// TIA Portal project "Project2_Pompe" (V15.1)

(* hardware
DEVICE "S71500/ET200MP station_1"  S7-1500 station
   slot 0: "Rail_0"  Rack  6ES7 590-1***0-0AA0
   slot 1: "PLC_1"  CPU 1513-1 PN  6ES7 513-1AL02-0AB0  V2.6
      slot 3: "CPU display_1"  6ES7591-1AA00-0AA0
DEVICE "HMI_1"  KTP900 Basic PN
   slot 0: "HMI_1"  KTP900 Basic PN  6AV2 123-2JB03-0AX0  15.1.0.0
   slot 1: "HMI_RT_1"  KTP900 Basic PN  6AV2 123-2JB03-0AX0  15.1.0.0
   slot 5: "HMI_1.IE_CP_1"  PROFINET Interface  15.0.1.0
      slot 1: "PROFINET Interface_1"  PROFINET Interface
         slot 1: "Port_1"  Port
*)

// ===== PLC "PLC_1"  CPU 1513-1 PN =====

VAR_GLOBAL   // PLC tag table "Default tag table"
   "Clock_Byte" AT %MB0 : Byte;
   "Clock_10Hz" AT %M0.0 : Bool;
   "Clock_5Hz" AT %M0.1 : Bool;
   "Clock_2.5Hz" AT %M0.2 : Bool;
   "Clock_2Hz" AT %M0.3 : Bool;
   "Clock_1.25Hz" AT %M0.4 : Bool;
   "Clock_1Hz" AT %M0.5 : Bool;
   "Clock_0.625Hz" AT %M0.6 : Bool;
   "Clock_0.5Hz" AT %M0.7 : Bool;
END_VAR

VAR_GLOBAL   // PLC tag table "Intrari"
   "S1(clk)" AT %I0.0 : Bool;
   "S2(ctrclk)" AT %I0.1 : Bool;
   "s0(stop)" AT %I0.2 : Bool;
   "ptc(esd)" AT %I0.3 : Bool;
   "ss" AT %I0.4 : Bool;
END_VAR

VAR_GLOBAL   // PLC tag table "Iesiri"
   "K1(clk)" AT %Q0.0 : Bool;
   "K2(ctrclk)" AT %Q0.1 : Bool;
   "K3(triunghi)" AT %Q0.2 : Bool;
   "K4(stea)" AT %Q0.3 : Bool;
END_VAR

VAR_GLOBAL   // PLC tag table "Auxiliare"
   "M_pornit" AT %M1.0 : Bool;
   "passed_k3" AT %M1.1 : Bool;
   "reset urgenta" AT %M1.2 : Bool;
   "temporizare K4" AT %M1.3 : Bool;
   "permisie start" AT %M1.4 : Bool;
   "urgenta bit" AT %M1.5 : Bool;
END_VAR

// folder: System blocks/Program resources

DATA_BLOCK "IEC_Timer_0_DB"   // DB1
{ S7_Optimized_Access := 'TRUE' }
AUTHOR : Simatic
FAMILY : IEC
NAME : IEC_TMR
VERSION : 1.0
// stored: InstanceOfName IEC_TIMER
"IEC_TIMER"
BEGIN
END_DATA_BLOCK

DATA_BLOCK "IEC_Timer_0_DB_1"   // DB2
{ S7_Optimized_Access := 'TRUE' }
AUTHOR : Simatic
FAMILY : IEC
NAME : IEC_TMR
VERSION : 1.0
// stored: InstanceOfName IEC_TIMER
"IEC_TIMER"
BEGIN
END_DATA_BLOCK

// folder: (top level)

FUNCTION_BLOCK "Block_1"   // FB1, LAD
{ S7_Optimized_Access := 'TRUE' }
VERSION : 0.1
   VAR_INPUT
      start : Bool;
      stop : Bool;
      ESD : Bool;
   END_VAR
   VAR_OUTPUT
      "comanda motor" : Bool;
   END_VAR
BEGIN

REGION Network 1
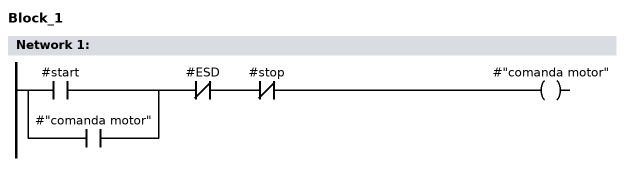
   RUNG wire#powerrail
      Contact( #start )
      wire#w1
      I_Contact( #ESD )
      I_Contact( #stop )
      Coil( #"comanda motor" )
   END_RUNG
   RUNG wire#powerrail
      Contact( #"comanda motor" )
   END_RUNG wire#w1
   // the same network as SCL:
   #"comanda motor" := (#start OR #"comanda motor") AND NOT #ESD AND NOT #stop;
END_REGION
END_FUNCTION_BLOCK

ORGANIZATION_BLOCK "Main"   // OB1, LAD, ProgramCycle
TITLE = "Main Program Sweep (Cycle)"
{ S7_Optimized_Access := 'TRUE' }
VERSION : 0.1
   VAR_INPUT
      Initial_Call : Bool;   // Initial call of this OB
      Remanence : Bool;   // =True, if remanent data are available
   END_VAR
BEGIN

REGION Network 1: selecteaza pe ce directie sa porneasca
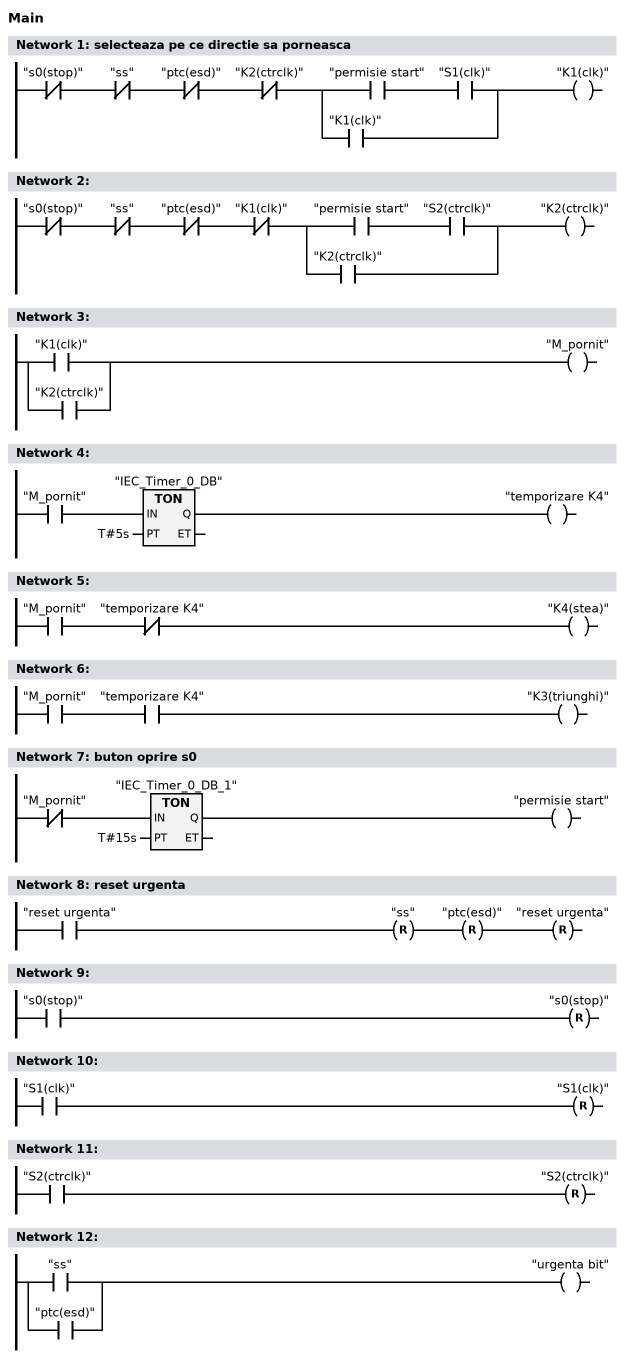
   RUNG wire#powerrail
      I_Contact( "s0(stop)" )
      I_Contact( "ss" )
      I_Contact( "ptc(esd)" )
      I_Contact( "K2(ctrclk)" )
      wire#w1
      Contact( "permisie start" )
      Contact( "S1(clk)" )
      wire#w2
      Coil( "K1(clk)" )
   END_RUNG
   RUNG wire#w1
      Contact( "K1(clk)" )
   END_RUNG wire#w2
   // the same network as SCL:
   "K1(clk)" := NOT "s0(stop)" AND NOT "ss" AND NOT "ptc(esd)" AND NOT "K2(ctrclk)" AND (("permisie start" AND "S1(clk)") OR "K1(clk)");
END_REGION

REGION Network 2
   RUNG wire#powerrail
      I_Contact( "s0(stop)" )
      I_Contact( "ss" )
      I_Contact( "ptc(esd)" )
      I_Contact( "K1(clk)" )
      wire#w1
      Contact( "permisie start" )
      Contact( "S2(ctrclk)" )
      wire#w2
      Coil( "K2(ctrclk)" )
   END_RUNG
   RUNG wire#w1
      Contact( "K2(ctrclk)" )
   END_RUNG wire#w2
   // the same network as SCL:
   "K2(ctrclk)" := NOT "s0(stop)" AND NOT "ss" AND NOT "ptc(esd)" AND NOT "K1(clk)" AND (("permisie start" AND "S2(ctrclk)") OR "K2(ctrclk)");
END_REGION

REGION Network 3
   RUNG wire#powerrail
      Contact( "K1(clk)" )
      wire#w1
      Coil( "M_pornit" )
   END_RUNG
   RUNG wire#powerrail
      Contact( "K2(ctrclk)" )
   END_RUNG wire#w1
   // the same network as SCL:
   "M_pornit" := "K1(clk)" OR "K2(ctrclk)";
END_REGION

REGION Network 4
   "IEC_Timer_0_DB".TON(IN := "M_pornit", PT := T#5s);
   "temporizare K4" := "IEC_Timer_0_DB".Q;
END_REGION

REGION Network 5
   RUNG wire#powerrail
      Contact( "M_pornit" )
      I_Contact( "temporizare K4" )
      Coil( "K4(stea)" )
   END_RUNG
   // the same network as SCL:
   "K4(stea)" := "M_pornit" AND NOT "temporizare K4";
END_REGION

REGION Network 6
   RUNG wire#powerrail
      Contact( "M_pornit" )
      Contact( "temporizare K4" )
      Coil( "K3(triunghi)" )
   END_RUNG
   // the same network as SCL:
   "K3(triunghi)" := "M_pornit" AND "temporizare K4";
END_REGION

REGION Network 7: buton oprire s0
   "IEC_Timer_0_DB_1".TON(IN := NOT "M_pornit", PT := T#15s);
   "permisie start" := "IEC_Timer_0_DB_1".Q;
END_REGION

REGION Network 8: reset urgenta
   RUNG wire#powerrail
      Contact( "reset urgenta" )
      R_Coil( "ss" )
      R_Coil( "ptc(esd)" )
      R_Coil( "reset urgenta" )
   END_RUNG
   // the same network as SCL:
   IF "reset urgenta" THEN
       "ss" := FALSE;
       "ptc(esd)" := FALSE;
       "reset urgenta" := FALSE;
   END_IF;
END_REGION

REGION Network 9
   RUNG wire#powerrail
      Contact( "s0(stop)" )
      R_Coil( "s0(stop)" )
   END_RUNG
   // the same network as SCL:
   IF "s0(stop)" THEN "s0(stop)" := FALSE; END_IF;
END_REGION

REGION Network 10
   RUNG wire#powerrail
      Contact( "S1(clk)" )
      R_Coil( "S1(clk)" )
   END_RUNG
   // the same network as SCL:
   IF "S1(clk)" THEN "S1(clk)" := FALSE; END_IF;
END_REGION

REGION Network 11
   RUNG wire#powerrail
      Contact( "S2(ctrclk)" )
      R_Coil( "S2(ctrclk)" )
   END_RUNG
   // the same network as SCL:
   IF "S2(ctrclk)" THEN "S2(ctrclk)" := FALSE; END_IF;
END_REGION

REGION Network 12
   RUNG wire#powerrail
      Contact( "ss" )
      wire#w1
      Coil( "urgenta bit" )
   END_RUNG
   RUNG wire#powerrail
      Contact( "ptc(esd)" )
   END_RUNG wire#w1
   // the same network as SCL:
   "urgenta bit" := "ss" OR "ptc(esd)";
END_REGION
END_ORGANIZATION_BLOCK

(* ===== HMI "HMI_RT_1" =====
system functions are stored by id; their names below are inferred from use
connection "HMI_Connection_1": ETHERNET, SMART_S7_1500_OMS

HMI tags "Default tag table"
   "Tag_ScreenNumber" : UInt, internal
   "s0(stop)" : Bool = PLC "s0(stop)" AT %I0.2, 1 s
   "S1(clk)" : Bool = PLC "S1(clk)" AT %I0.0, 1 s
   "S2(ctrclk)" : Bool = PLC "S2(ctrclk)" AT %I0.1, 1 s
   "IEC_Timer_0_DB_1_ET" : Time = PLC IEC_Timer_0_DB_1.ET, 1 s
   "IEC_Timer_0_DB_ET" : Time = PLC IEC_Timer_0_DB.ET, 1 s
   "K1(clk)" : Bool = PLC "K1(clk)" AT %Q0.0, 1 s
   "K2(ctrclk)" : Bool = PLC "K2(ctrclk)" AT %Q0.1, 1 s
   "K3(triunghi)" : Bool = PLC "K3(triunghi)" AT %Q0.2, 1 s
   "K4(stea)" : Bool = PLC "K4(stea)" AT %Q0.3, 1 s
   "ss" : Bool = PLC ss AT %I0.4, 1 s
   "M_pornit" : Bool = PLC M_pornit AT %M1.0, 1 s
   "reset urgenta" : Bool = PLC "reset urgenta" AT %M1.2, 1 s
   "ptc(esd)" : Bool = PLC "ptc(esd)" AT %I0.3, 1 s
   "urgenta bit" : Bool = PLC "urgenta bit" AT %M1.5, 1 s

Template "Template_1" 800x480
   Button "Exit" at 722,440 size 55x39; TextOff 'Exit'; PictureOff "ExitRuntime_KTP900_Basic_PN_TR"; PictureOn "ExitRuntime_KTP900_Basic_PN_TR"
      on Release: StopRuntime(0)
   Button "Template_Button" at 622,440 size 55x39; TextOff 'Text'
   Button "Template_Button_1" at 522,440 size 55x39; TextOff 'Text'
   Button "Template_Button_2" at 422,440 size 55x39; TextOff 'Text'
   Button "Template_Button_3" at 322,440 size 55x39; TextOff 'Text'
   Button "Template_Button_4" at 222,440 size 55x39; TextOff 'Text'
   Button "Alarms" at 122,440 size 55x39; TextOff 'Alarms'; PictureOff "AlarmDisplay_KTP900_Basic_PN_TR"; PictureOn "AlarmDisplay_KTP900_Basic_PN_TR"
      on Release: function_ef3f5d25("Alarm window_Unacknowledged", -1)
   Button "Start screen" at 22,440 size 55x39; TextOff 'Start screen'; PictureOff "NavigateHome_KTP900_Basic_PN_TR"; PictureOn "NavigateHome_KTP900_Basic_PN_TR"
      on Release: ActivateScreen("Root screen", 0)
   SymbolicIOField "Symbolic_IO_Field_Screen" at 73,7 size 620x26; TextOff '0'; TextOn '1'; TextList "TextList_ScreenNames"
      ProcessValue <- "Tag_ScreenNumber"
      on Change: ActivateScreenByNumber("Tag_ScreenNumber", 0)
   DateTimeField "HmiScreenItemData" at 695,20 size 105x20
   DateTimeField "HmiScreenItemData_1" at 695,0 size 105x20
   GraphicView "Logo" at 0,0 size 71x40; Picture "Logo of HMI_1"

screen "Root screen" 800x480, template "Template_1"
   on GenerateScreen: SetTag("Tag_ScreenNumber", 1)
   Circle "Circle_1" at 129,113 size 86x86
      Appearance <- "M_pornit"
   Group "Group" at 129,113 size 89x87
   TextField "Text field_1" at 156,61 size 35x20; Text 'Stop'
   TextField "Text field_2" at 18,64 size 67x20; Text 'Clockwise'
   TextField "Text field_3" at 256,66 size 87x20; Text 'CtrClockwise'
   Button "Button_1" at 657,68 size 96x32; TextOff 'Stop'
      on Click: SetBit("s0(stop)")
   TextField "Text field_4" at 619,73 size 21x20; Text 'S0'
   Button "Button_2" at 658,118 size 96x32; TextOff 'Start K1'
      on Click: SetBit("S1(clk)")
   Button "Button_3" at 658,167 size 96x32; TextOff 'Start K2'
      on Click: SetBit("S2(ctrclk)")
   Circle "Circle_3" at 606,113 size 42x42
      Appearance <- "K1(clk)"
   Circle "Circle_4" at 606,168 size 42x42
      Appearance <- "K2(ctrclk)"
   TextField "Text field_5" at 570,122 size 21x20; Text 'S1'
   TextField "Text field_6" at 570,175 size 21x20; Text 'S2'
   Button "Button_4" at 623,351 size 96x32; TextOff 'ESD'
      on Click: SetBit("ss")
   TextField "Text field_7" at 584,353 size 21x20; Text 'SS'
   Circle "Circle_2" at 331,307 size 79x79
      Appearance <- "K3(triunghi)"
   Circle "Circle_5" at 440,306 size 79x79
      Appearance <- "K4(stea)"
   TextField "Text field_8" at 362,334 size 21x20; Text 'K3'
   TextField "Text field_9" at 473,336 size 21x20; Text 'K4'
   Button "Button_5" at 21,390 size 96x32; TextOff 'Just press'
   Button "Button_6" at 623,397 size 96x32; TextOff 'Reset ESD'
      on Click: SetBit("reset urgenta")
   IOField "I/O field_1" at 526,71 size 44x32; FormatPattern 99; Unit s
      ProcessValue <- "IEC_Timer_0_DB_1_ET"
   IOField "I/O field_2" at 458,259 size 56x32; FormatPattern 999; Unit s
      ProcessValue <- "IEC_Timer_0_DB_ET"
   TextField "Text field_10" at 453,239 size 60x20; Text 'Timer K4'
   TextField "Text field_11" at 505,51 size 92x20; Text 'Timer to Stop'
   Circle "Circle_6" at 128,271 size 101x101
      Appearance <- "M_pornit"
   TextField "Text field_12" at 73,307 size 44x20; Text 'Motor'
   Group "Group_1" at 262,108 size 89x87
   Group "Group_2" at 17,114 size 89x87
   Ellipse "Ellipse_1" at 640,317 size 67x28
      Appearance <- "urgenta bit"
   Circle "Circle_7" at 262,108 size 86x86
      Appearance <- "K2(ctrclk)"
   Circle "Circle_8" at 17,114 size 86x86
      Appearance <- "K1(clk)"
*)